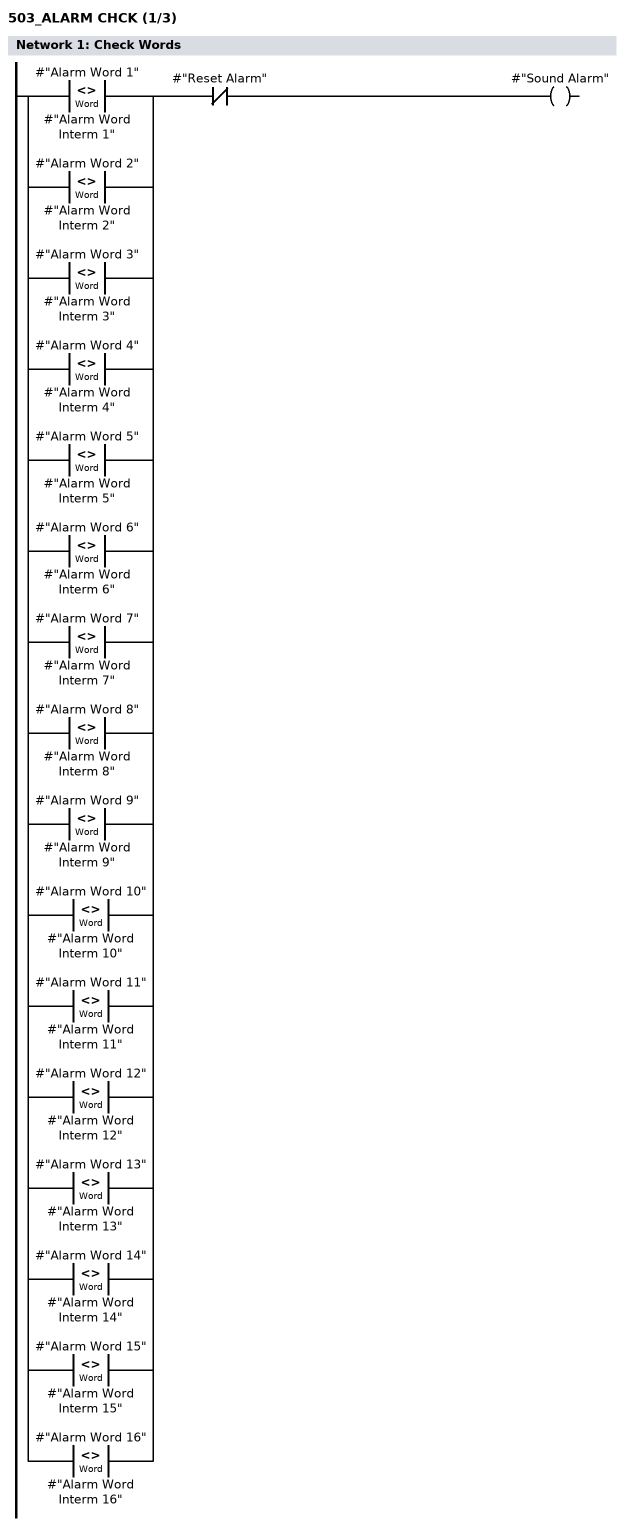
   RUNG wire#powerrail
      { S7_Templates := "SrcType := Word" } NE_Contact(in1 := #"Alarm Word 1", in2 := #"Alarm Word Interm 1")
      wire#w1
      I_Contact( #"Reset Alarm" )
      Coil( #"Sound Alarm" )
   END_RUNG
   RUNG wire#powerrail
      { S7_Templates := "SrcType := Word" } NE_Contact(in1 := #"Alarm Word 2", in2 := #"Alarm Word Interm 2")
   END_RUNG wire#w1
   RUNG wire#powerrail
      { S7_Templates := "SrcType := Word" } NE_Contact(in1 := #"Alarm Word 3", in2 := #"Alarm Word Interm 3")
   END_RUNG wire#w1
   RUNG wire#powerrail
      { S7_Templates := "SrcType := Word" } NE_Contact(in1 := #"Alarm Word 4", in2 := #"Alarm Word Interm 4")
   END_RUNG wire#w1
   RUNG wire#powerrail
      { S7_Templates := "SrcType := Word" } NE_Contact(in1 := #"Alarm Word 5", in2 := #"Alarm Word Interm 5")
   END_RUNG wire#w1
   RUNG wire#powerrail
      { S7_Templates := "SrcType := Word" } NE_Contact(in1 := #"Alarm Word 6", in2 := #"Alarm Word Interm 6")
   END_RUNG wire#w1
   RUNG wire#powerrail
      { S7_Templates := "SrcType := Word" } NE_Contact(in1 := #"Alarm Word 7", in2 := #"Alarm Word Interm 7")
   END_RUNG wire#w1
   RUNG wire#powerrail
      { S7_Templates := "SrcType := Word" } NE_Contact(in1 := #"Alarm Word 8", in2 := #"Alarm Word Interm 8")
   END_RUNG wire#w1
   RUNG wire#powerrail
      { S7_Templates := "SrcType := Word" } NE_Contact(in1 := #"Alarm Word 9", in2 := #"Alarm Word Interm 9")
   END_RUNG wire#w1
   RUNG wire#powerrail
      { S7_Templates := "SrcType := Word" } NE_Contact(in1 := #"Alarm Word 10", in2 := #"Alarm Word Interm 10")
   END_RUNG wire#w1
   RUNG wire#powerrail
      { S7_Templates := "SrcType := Word" } NE_Contact(in1 := #"Alarm Word 11", in2 := #"Alarm Word Interm 11")
   END_RUNG wire#w1
   RUNG wire#powerrail
      { S7_Templates := "SrcType := Word" } NE_Contact(in1 := #"Alarm Word 12", in2 := #"Alarm Word Interm 12")
   END_RUNG wire#w1
   RUNG wire#powerrail
      { S7_Templates := "SrcType := Word" } NE_Contact(in1 := #"Alarm Word 13", in2 := #"Alarm Word Interm 13")
   END_RUNG wire#w1
   RUNG wire#powerrail
      { S7_Templates := "SrcType := Word" } NE_Contact(in1 := #"Alarm Word 14", in2 := #"Alarm Word Interm 14")
   END_RUNG wire#w1
   RUNG wire#powerrail
      { S7_Templates := "SrcType := Word" } NE_Contact(in1 := #"Alarm Word 15", in2 := #"Alarm Word Interm 15")
   END_RUNG wire#w1
   RUNG wire#powerrail
      { S7_Templates := "SrcType := Word" } NE_Contact(in1 := #"Alarm Word 16", in2 := #"Alarm Word Interm 16")
   END_RUNG wire#w1
   // the same network as SCL:
   #"Sound Alarm" := ((#"Alarm Word 1" <> #"Alarm Word Interm 1") OR (#"Alarm Word 2" <> #"Alarm Word Interm 2") OR (#"Alarm Word 3" <> #"Alarm Word Interm 3") OR (#"Alarm Word 4" <> #"Alarm Word Interm 4") OR (#"Alarm Word 5" <> #"Alarm Word Interm 5") OR (#"Alarm Word 6" <> #"Alarm Word Interm 6") OR (#"Alarm Word 7" <> #"Alarm Word Interm 7") OR (#"Alarm Word 8" <> #"Alarm Word Interm 8") OR (#"Alarm Word 9" <> #"Alarm Word Interm 9") OR (#"Alarm Word 10" <> #"Alarm Word Interm 10") OR (#"Alarm Word 11" <> #"Alarm Word Interm 11") OR (#"Alarm Word 12" <> #"Alarm Word Interm 12") OR (#"Alarm Word 13" <> #"Alarm Word Interm 13") OR (#"Alarm Word 14" <> #"Alarm Word Interm 14") OR (#"Alarm Word 15" <> #"Alarm Word Interm 15") OR (#"Alarm Word 16" <> #"Alarm Word Interm 16")) AND NOT #"Reset Alarm";
END_REGION

REGION Network 2
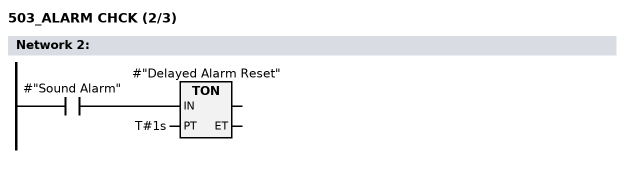
   #"Delayed Alarm Reset"(IN := #"Sound Alarm", PT := T#1s);   // TON
END_REGION

REGION Network 3: Move Words
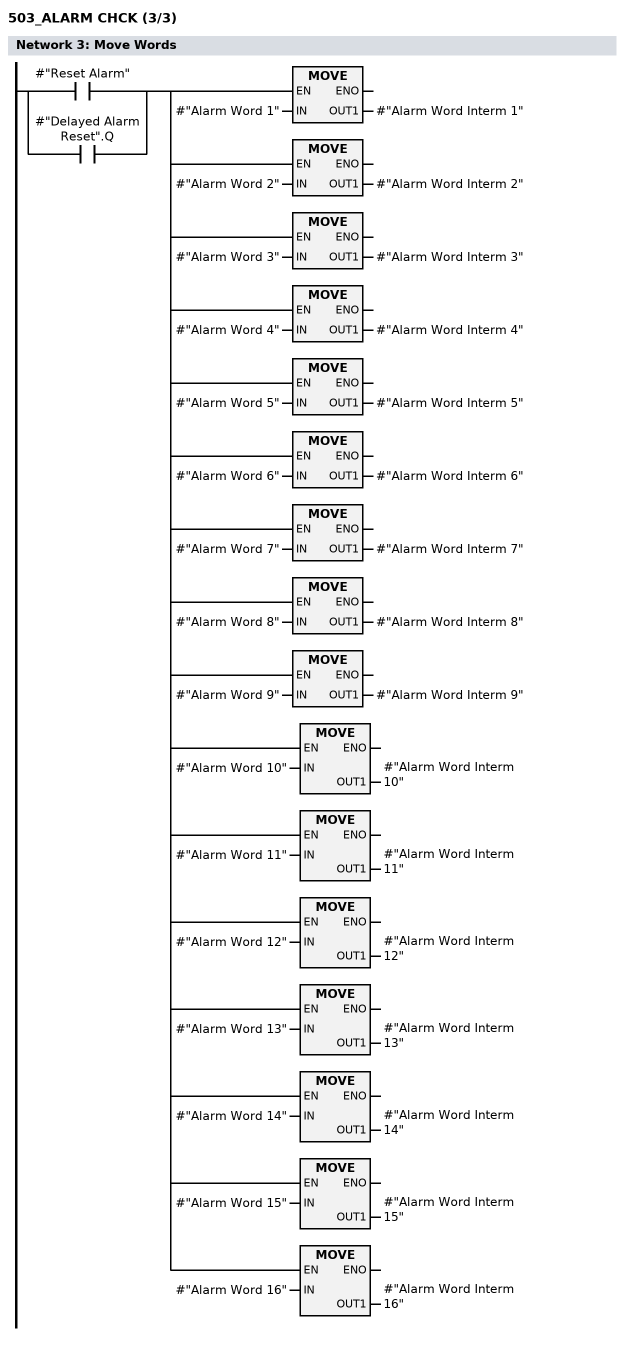
   RUNG wire#powerrail
      Contact( #"Reset Alarm" )
      wire#w1
      Move(in := #"Alarm Word 1", out1 => #"Alarm Word Interm 1")
   END_RUNG
   RUNG wire#powerrail
      Contact( #"Delayed Alarm Reset".Q )
   END_RUNG wire#w1
   RUNG wire#w1
      Move(in := #"Alarm Word 2", out1 => #"Alarm Word Interm 2")
   END_RUNG
   RUNG wire#w1
      Move(in := #"Alarm Word 3", out1 => #"Alarm Word Interm 3")
   END_RUNG
   RUNG wire#w1
      Move(in := #"Alarm Word 4", out1 => #"Alarm Word Interm 4")
   END_RUNG
   RUNG wire#w1
      Move(in := #"Alarm Word 5", out1 => #"Alarm Word Interm 5")
   END_RUNG
   RUNG wire#w1
      Move(in := #"Alarm Word 6", out1 => #"Alarm Word Interm 6")
   END_RUNG
   RUNG wire#w1
      Move(in := #"Alarm Word 7", out1 => #"Alarm Word Interm 7")
   END_RUNG
   RUNG wire#w1
      Move(in := #"Alarm Word 8", out1 => #"Alarm Word Interm 8")
   END_RUNG
   RUNG wire#w1
      Move(in := #"Alarm Word 9", out1 => #"Alarm Word Interm 9")
   END_RUNG
   RUNG wire#w1
      Move(in := #"Alarm Word 10", out1 => #"Alarm Word Interm 10")
   END_RUNG
   RUNG wire#w1
      Move(in := #"Alarm Word 11", out1 => #"Alarm Word Interm 11")
   END_RUNG
   RUNG wire#w1
      Move(in := #"Alarm Word 12", out1 => #"Alarm Word Interm 12")
   END_RUNG
   RUNG wire#w1
      Move(in := #"Alarm Word 13", out1 => #"Alarm Word Interm 13")
   END_RUNG
   RUNG wire#w1
      Move(in := #"Alarm Word 14", out1 => #"Alarm Word Interm 14")
   END_RUNG
   RUNG wire#w1
      Move(in := #"Alarm Word 15", out1 => #"Alarm Word Interm 15")
   END_RUNG
   RUNG wire#w1
      Move(in := #"Alarm Word 16", out1 => #"Alarm Word Interm 16")
   END_RUNG
   // the same network as SCL:
   IF #"Reset Alarm" OR #"Delayed Alarm Reset".Q THEN
       #"Alarm Word Interm 1" := #"Alarm Word 1";
       #"Alarm Word Interm 2" := #"Alarm Word 2";
       #"Alarm Word Interm 3" := #"Alarm Word 3";
       #"Alarm Word Interm 4" := #"Alarm Word 4";
       #"Alarm Word Interm 5" := #"Alarm Word 5";
       #"Alarm Word Interm 6" := #"Alarm Word 6";
       #"Alarm Word Interm 7" := #"Alarm Word 7";
       #"Alarm Word Interm 8" := #"Alarm Word 8";
       #"Alarm Word Interm 9" := #"Alarm Word 9";
       #"Alarm Word Interm 10" := #"Alarm Word 10";
       #"Alarm Word Interm 11" := #"Alarm Word 11";
       #"Alarm Word Interm 12" := #"Alarm Word 12";
       #"Alarm Word Interm 13" := #"Alarm Word 13";
       #"Alarm Word Interm 14" := #"Alarm Word 14";
       #"Alarm Word Interm 15" := #"Alarm Word 15";
       #"Alarm Word Interm 16" := #"Alarm Word 16";
   END_IF;
END_REGION
END_FUNCTION_BLOCK

FUNCTION_BLOCK "Choose"   // FB509, LAD
{ S7_Optimized_Access := 'TRUE' }
VERSION : 0.1
   VAR_INPUT
      Choose : Bool;
      "Option 1" : DInt;
      "Option 2" : DInt;
   END_VAR
   VAR_OUTPUT
      Output : DInt;
   END_VAR
   VAR
      True : Bool;
      False : Bool;
      "Option 1 M" : DInt;
      "Option 2 M" : DInt;
      "Choose Internal" : Bool;
      "Puls Aux" : Struct
         "Puls Aux 1" : Bool;
         "Puls Aux 2" : Bool;
         "Puls Aux 3" : Bool;
         "Puls Aux 4" : Bool;
         "Puls Aux 5" : Bool;
         "Puls Aux 6" : Bool;
      END_STRUCT;
      "TP P CHOOSE1" : TP_TIME;
      "TP N CHOOSE2" : TP_TIME;
      "TP N CHOOSE1" : TP_TIME;
      "TP P CHOOSE2" : TP_TIME;
      R_TRIG_Instance : R_TRIG;
      Puls : TP_TIME;
   END_VAR
   VAR_TEMP   // added for the SCL form of the ladder/FBD networks
      _w1 : Bool;
      _w2 : Bool;
      _w3 : Bool;
      _w4 : Bool;
   END_VAR
BEGIN

REGION Network 1: False/True
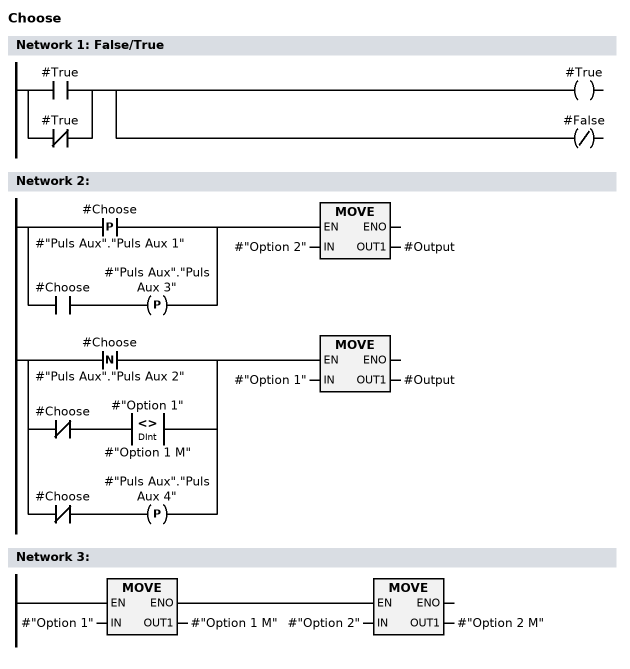
   RUNG wire#powerrail
      Contact( #True )
      wire#w1
      Coil( #True )
   END_RUNG
   RUNG wire#powerrail
      I_Contact( #True )
   END_RUNG wire#w1
   RUNG wire#w1
      I_Coil( #False )
   END_RUNG
   // the same network as SCL:
   #True := #True OR NOT #True;
   #False := NOT #True;
END_REGION

REGION Network 2
   RUNG wire#powerrail
      P_Contact(operand := #Choose, bit := #"Puls Aux"."Puls Aux 1")
      wire#w1
      Move(in := #"Option 2", out1 => #Output)
   END_RUNG
   RUNG wire#powerrail
      Contact( #Choose )
      P_Trig( #"Puls Aux"."Puls Aux 3" )
   END_RUNG wire#w1
   RUNG wire#powerrail
      N_Contact(operand := #Choose, bit := #"Puls Aux"."Puls Aux 2")
      wire#w2
      Move(in := #"Option 1", out1 => #Output)
   END_RUNG
   RUNG wire#powerrail
      I_Contact( #Choose )
      { S7_Templates := "SrcType := DInt" } NE_Contact(in1 := #"Option 1", in2 := #"Option 1 M")
   END_RUNG wire#w2
   RUNG wire#powerrail
      I_Contact( #Choose )
      P_Trig( #"Puls Aux"."Puls Aux 4" )
   END_RUNG wire#w2
   // the same network as SCL:
   #_w1 := #Choose AND NOT #"Puls Aux"."Puls Aux 1";   // rising edge of #Choose
   #"Puls Aux"."Puls Aux 1" := #Choose;
   #_w2 := #Choose AND NOT #"Puls Aux"."Puls Aux 3";   // rising edge
   #"Puls Aux"."Puls Aux 3" := #Choose;
   IF #_w1 OR #_w2 THEN #Output := #"Option 2"; END_IF;
   #_w3 := NOT #Choose AND #"Puls Aux"."Puls Aux 2";   // falling edge of #Choose
   #"Puls Aux"."Puls Aux 2" := #Choose;
   #_w4 := NOT #Choose AND NOT #"Puls Aux"."Puls Aux 4";   // rising edge
   #"Puls Aux"."Puls Aux 4" := NOT #Choose;
   IF #_w3 OR (NOT #Choose AND (#"Option 1" <> #"Option 1 M")) OR #_w4 THEN #Output := #"Option 1"; END_IF;
END_REGION

REGION Network 3
   RUNG wire#powerrail
      Move(in := #"Option 1", out1 => #"Option 1 M")
      Move(in := #"Option 2", out1 => #"Option 2 M")
   END_RUNG
   // the same network as SCL:
   #"Option 1 M" := #"Option 1";
   #"Option 2 M" := #"Option 2";
END_REGION
END_FUNCTION_BLOCK

FUNCTION_BLOCK "Flip Flop"   // FB510, LAD
{ S7_Optimized_Access := 'TRUE' }
VERSION : 0.1
   VAR_INPUT
      Input : Bool;
   END_VAR
   VAR_OUTPUT
      Output : Bool;
   END_VAR
   VAR
      SetOutputFlag : Bool;
   END_VAR
   VAR_TEMP   // added for the SCL form of the ladder/FBD networks
      _w1 : Bool;
      _w2 : Bool;
   END_VAR
BEGIN

REGION Network 2: Set Group SR
   // HMI Button to be set as SetTagWhileKeyPres
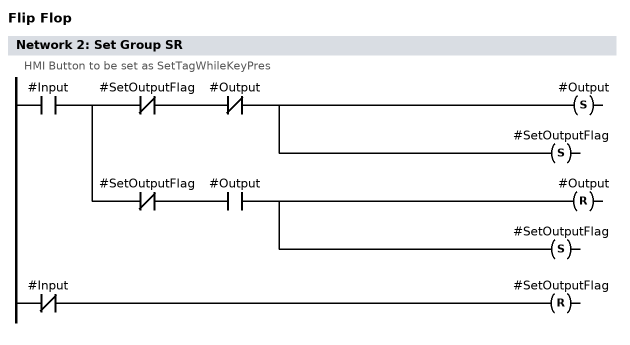
   RUNG wire#powerrail
      Contact( #Input )
      wire#w1
      I_Contact( #SetOutputFlag )
      I_Contact( #Output )
      wire#w2
      S_Coil( #Output )
   END_RUNG
   RUNG wire#w2
      S_Coil( #SetOutputFlag )
   END_RUNG
   RUNG wire#w1
      I_Contact( #SetOutputFlag )
      Contact( #Output )
      wire#w3
      R_Coil( #Output )
   END_RUNG
   RUNG wire#w3
      S_Coil( #SetOutputFlag )
   END_RUNG
   RUNG wire#powerrail
      I_Contact( #Input )
      R_Coil( #SetOutputFlag )
   END_RUNG
   // the same network as SCL:
   #_w1 := #Input AND NOT #SetOutputFlag AND NOT #Output;
   IF #_w1 THEN
       #Output := TRUE;
       #SetOutputFlag := TRUE;
   END_IF;
   #_w2 := #Input AND NOT #SetOutputFlag AND #Output;
   IF #_w2 THEN
       #Output := FALSE;
       #SetOutputFlag := TRUE;
   END_IF;
   IF NOT #Input THEN #SetOutputFlag := FALSE; END_IF;
END_REGION
END_FUNCTION_BLOCK

FUNCTION_BLOCK "Memory"   // FB511, LAD
{ S7_Optimized_Access := 'TRUE' }
VERSION : 0.1
   VAR_INPUT
      Enable : Bool;
      Negated : Bool := true;
      "Memorise/Remember" : Bool;
      Value : Int;
   END_VAR
   VAR_OUTPUT
      Remember : Int;
   END_VAR
   VAR RETAIN
      Memory : Int;
   END_VAR
   VAR
      PulsAuxP : Bool;
      PulsAuxN : Bool;
      SetOutputFlag : Bool;
      Output : Bool;
   END_VAR
   VAR_TEMP   // added for the SCL form of the ladder/FBD networks
      _w1 : Bool;
      _w2 : Bool;
      _w3 : Bool;
   END_VAR
BEGIN

REGION Network 1: Set Group SR
   // HMI Button to be set as SetTagWhileKeyPres
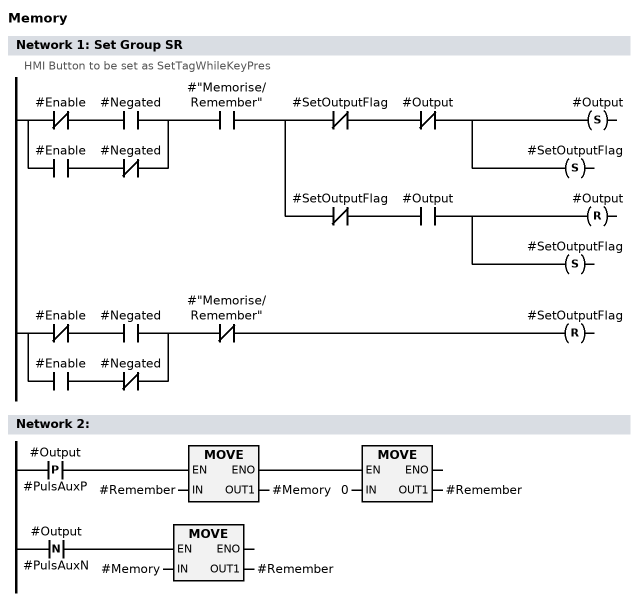
   RUNG wire#powerrail
      I_Contact( #Enable )
      Contact( #Negated )
      wire#w1
      Contact( #"Memorise/Remember" )
      wire#w2
      I_Contact( #SetOutputFlag )
      I_Contact( #Output )
      wire#w3
      S_Coil( #Output )
   END_RUNG
   RUNG wire#powerrail
      Contact( #Enable )
      I_Contact( #Negated )
   END_RUNG wire#w1
   RUNG wire#w3
      S_Coil( #SetOutputFlag )
   END_RUNG
   RUNG wire#w2
      I_Contact( #SetOutputFlag )
      Contact( #Output )
      wire#w4
      R_Coil( #Output )
   END_RUNG
   RUNG wire#w4
      S_Coil( #SetOutputFlag )
   END_RUNG
   RUNG wire#powerrail
      I_Contact( #Enable )
      Contact( #Negated )
      wire#w5
      I_Contact( #"Memorise/Remember" )
      R_Coil( #SetOutputFlag )
   END_RUNG
   RUNG wire#powerrail
      Contact( #Enable )
      I_Contact( #Negated )
   END_RUNG wire#w5
   // the same network as SCL:
   #_w1 := ((NOT #Enable AND #Negated) OR (#Enable AND NOT #Negated)) AND #"Memorise/Remember";
   #_w2 := #_w1 AND NOT #SetOutputFlag AND NOT #Output;
   IF #_w2 THEN
       #Output := TRUE;
       #SetOutputFlag := TRUE;
   END_IF;
   #_w3 := #_w1 AND NOT #SetOutputFlag AND #Output;
   IF #_w3 THEN
       #Output := FALSE;
       #SetOutputFlag := TRUE;
   END_IF;
   IF ((NOT #Enable AND #Negated) OR (#Enable AND NOT #Negated)) AND NOT #"Memorise/Remember" THEN
       #SetOutputFlag := FALSE;
   END_IF;
END_REGION

REGION Network 2
   RUNG wire#powerrail
      P_Contact(operand := #Output, bit := #PulsAuxP)
      Move(in := #Remember, out1 => #Memory)
      Move(in := 0, out1 => #Remember)
   END_RUNG
   RUNG wire#powerrail
      N_Contact(operand := #Output, bit := #PulsAuxN)
      Move(in := #Memory, out1 => #Remember)
   END_RUNG
   // the same network as SCL:
   #_w1 := #Output AND NOT #PulsAuxP;   // rising edge of #Output
   #PulsAuxP := #Output;
   IF #_w1 THEN
       #Memory := #Remember;
       #Remember := 0;
   END_IF;
   #_w2 := NOT #Output AND #PulsAuxN;   // falling edge of #Output
   #PulsAuxN := #Output;
   IF #_w2 THEN #Remember := #Memory; END_IF;
END_REGION
END_FUNCTION_BLOCK

FUNCTION_BLOCK "Sequence Times"   // FB512, LAD
{ S7_Optimized_Access := 'TRUE' }
VERSION : 0.1
   VAR_INPUT
      "Start Jurney" : Bool;
      "Start De-Ox" : Bool;
      "Start Dwell" : Bool;
      "Start Re-Ox" : Bool;
      "Start Post-Dwell" : Bool;
      "Jurney Time" : Real := 30.0;   // Days
      "Pre-Dwell Time" : Real := 1.0;   // Hours
      "De-Ox Time" : Real := 12.0;   // Hours
      "De-Ox SP Time" : Real := 1.0;   // Hours
      "De-Ox O2 Confirm" : Real := 1.0;   // Minutes
      "Dwell Time" : Real := 60.0;   // Hours
      "Re-Ox Time" : Real := 6.0;   // Hours
      "Post-Dwell Time" : Real := 12.0;   // Hours
      "Offset Treatment Time" : Real := 0.0;   // Hours
      "Offset Treatment Time Extend" : Real := 13.0;
      "Offset De-Ox Time Extend" : Real;
      "Offset Re-Ox Time Extend" : Real;
      "Time to IGG Start Warning" : DInt;   // Hours
      Continue : Bool;
      Boost : Bool;
   END_VAR
   VAR_OUTPUT
      "Times Valid" : Bool;
      "Warn to IGG Start" : Bool;
      "Warn to GCU Start" : Bool;   // Warning to start GCU at Re-Ox
      "Pre-Dwell Done" : Bool;
      "De-Ox Done" : Bool;
      "Dwell Done" : Bool;
      "Re-Ox Done" : Bool;
      "Post-Dwell Done" : Bool;
      "Pre-Dwell Time Corected" : Real;
      "Voiage Time Invalid" : Bool;
   END_VAR
   VAR
      "Extra Time" : Real;
      "Jurney Aux" : Time;
      "Pre-Dwell Aux" : Real;
      "Pre-Dwell Aux Memory" : Real;
   END_VAR
   VAR RETAIN
      "Pre-Dwell Memory h" : Real;
   END_VAR
   VAR
      "De-Ox Aux" : Real;
      "De-Ox Aux Memory" : Real;
   END_VAR
   VAR RETAIN
      "De-Ox Memory h" : Real;
   END_VAR
   VAR
      "Dwell Aux" : Real;
      "Dwell Aux Memory" : Real;
   END_VAR
   VAR RETAIN
      "Dwell Memory h" : Real;
   END_VAR
   VAR
      "Re-Ox Aux" : Real;
      "Re-Ox Aux Memory" : Real;
   END_VAR
   VAR RETAIN
      "Re-Ox Memory h" : Real;
   END_VAR
   VAR
      "Post-Dwell Aux" : Real;
      "Post-Dwell Aux Memory" : Real;
   END_VAR
   VAR RETAIN
      "Post-Dwell Memory h" : Real;
   END_VAR
   VAR
      True : Bool;
      False : Bool;
      "Pulse Continue" : Bool;
      IEC_Timer_0_Instance : TON_TIME;
      "Jurney Time FB" : "Days Timer";
      "Pre-Dwell Timer" : "Hours Timer";
      "Dwell Timer" : "Hours Timer";
      "Post-Dwell Timer" : "Hours Timer";
      "Puls Timer" : TON_TIME;
      "Puls TP" : TP_TIME;
      "Treatment Timer" : "Hours Timer";
      "De-Ox Timer" : "Hours Timer";
      "Re-Ox Timer" : "Hours Timer";
      "Jurney Timer" : "Hours Timer";
      "Offset Timer" : "Hours Timer";
      "Flip Flop_Pre-Dwell" : "Flip Flop";
      "Choose_Instance_Pre-Dwell" : "Choose Real";
      "Choose_Instance_De-Ox" : "Choose Real";
      Choose_Instance_Dwell : "Choose Real";
      "Choose_Instance_Re-Ox" : "Choose Real";
      "Choose_Instance_Post-Dwell" : "Choose Real";
   END_VAR
   VAR_TEMP   // added for the SCL form of the ladder/FBD networks
      _w1 : Bool;
   END_VAR
BEGIN

REGION Network 1
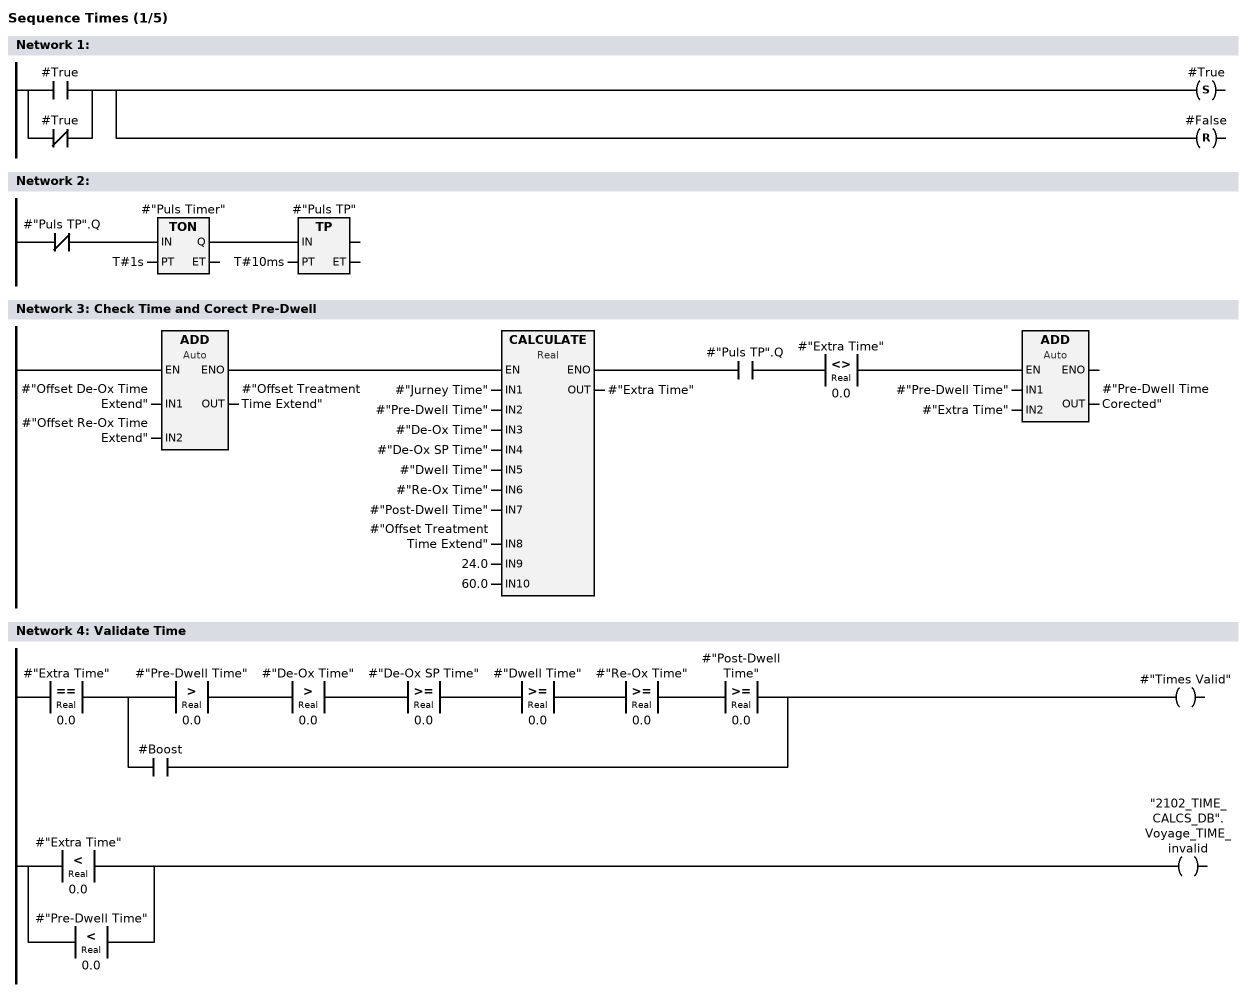
   RUNG wire#powerrail
      Contact( #True )
      wire#w1
      S_Coil( #True )
   END_RUNG
   RUNG wire#powerrail
      I_Contact( #True )
   END_RUNG wire#w1
   RUNG wire#w1
      R_Coil( #False )
   END_RUNG
   // the same network as SCL:
   #_w1 := #True OR NOT #True;
   IF #_w1 THEN
       #True := TRUE;
       #False := FALSE;
   END_IF;
END_REGION

REGION Network 2
   #"Puls Timer"(IN := NOT #"Puls TP".Q, PT := T#1s);   // TON
   #"Puls TP"(IN := #"Puls Timer".Q, PT := T#10ms);   // TP
END_REGION

REGION Network 3: Check Time and Corect Pre-Dwell
   RUNG wire#powerrail
      Add(in1 := #"Offset De-Ox Time Extend", in2 := #"Offset Re-Ox Time Extend", out => #"Offset Treatment Time Extend")
      { S7_Templates := "SrcType := Real"; S7_Expression := "IN1*IN9-(IN2+IN3+IN4+IN5+IN6+IN7+IN8)" } Calculate(in1 := #"Jurney Time", in2 := #"Pre-Dwell Time", in3 := #"De-Ox Time", in4 := #"De-Ox SP Time", in5 := #"Dwell Time", in6 := #"Re-Ox Time", in7 := #"Post-Dwell Time", in8 := #"Offset Treatment Time Extend", in9 := 24.0, in10 := 60.0, out => #"Extra Time")
      Contact( #"Puls TP".Q )
      { S7_Templates := "SrcType := Real" } NE_Contact(in1 := #"Extra Time", in2 := 0.0)
      Add(in1 := #"Pre-Dwell Time", in2 := #"Extra Time", out => #"Pre-Dwell Time Corected")
   END_RUNG
   // the same network as SCL:
   #"Offset Treatment Time Extend" := #"Offset De-Ox Time Extend" + #"Offset Re-Ox Time Extend";
   #"Extra Time" := #"Jurney Time"*24.0-(#"Pre-Dwell Time"+#"De-Ox Time"+#"De-Ox SP Time"+#"Dwell Time"+#"Re-Ox Time"+#"Post-Dwell Time"+#"Offset Treatment Time Extend");
   IF #"Puls TP".Q AND (#"Extra Time" <> 0.0) THEN
       #"Pre-Dwell Time Corected" := #"Pre-Dwell Time" + #"Extra Time";
   END_IF;
END_REGION

REGION Network 4: Validate Time
   RUNG wire#powerrail
      { S7_Templates := "SrcType := Real" } EQ_Contact(in1 := #"Extra Time", in2 := 0.0)
      wire#w1
      { S7_Templates := "SrcType := Real" } GT_Contact(in1 := #"Pre-Dwell Time", in2 := 0.0)
      { S7_Templates := "SrcType := Real" } GT_Contact(in1 := #"De-Ox Time", in2 := 0.0)
      { S7_Templates := "SrcType := Real" } GE_Contact(in1 := #"De-Ox SP Time", in2 := 0.0)
      { S7_Templates := "SrcType := Real" } GE_Contact(in1 := #"Dwell Time", in2 := 0.0)
      { S7_Templates := "SrcType := Real" } GE_Contact(in1 := #"Re-Ox Time", in2 := 0.0)
      { S7_Templates := "SrcType := Real" } GE_Contact(in1 := #"Post-Dwell Time", in2 := 0.0)
      wire#w2
      Coil( #"Times Valid" )
   END_RUNG
   RUNG wire#w1
      Contact( #Boost )
   END_RUNG wire#w2
   RUNG wire#powerrail
      { S7_Templates := "SrcType := Real" } LT_Contact(in1 := #"Extra Time", in2 := 0.0)
      wire#w3
      Coil( "2102_TIME_CALCS_DB".Voyage_TIME_invalid )
   END_RUNG
   RUNG wire#powerrail
      { S7_Templates := "SrcType := Real" } LT_Contact(in1 := #"Pre-Dwell Time", in2 := 0.0)
   END_RUNG wire#w3
   // the same network as SCL:
   #"Times Valid" := (#"Extra Time" = 0.0) AND (((#"Pre-Dwell Time" > 0.0) AND (#"De-Ox Time" > 0.0) AND (#"De-Ox SP Time" >= 0.0) AND (#"Dwell Time" >= 0.0) AND (#"Re-Ox Time" >= 0.0) AND (#"Post-Dwell Time" >= 0.0)) OR #Boost);
   "2102_TIME_CALCS_DB".Voyage_TIME_invalid := (#"Extra Time" < 0.0) OR (#"Pre-Dwell Time" < 0.0);
END_REGION

REGION Network 5: Total Sequence Time
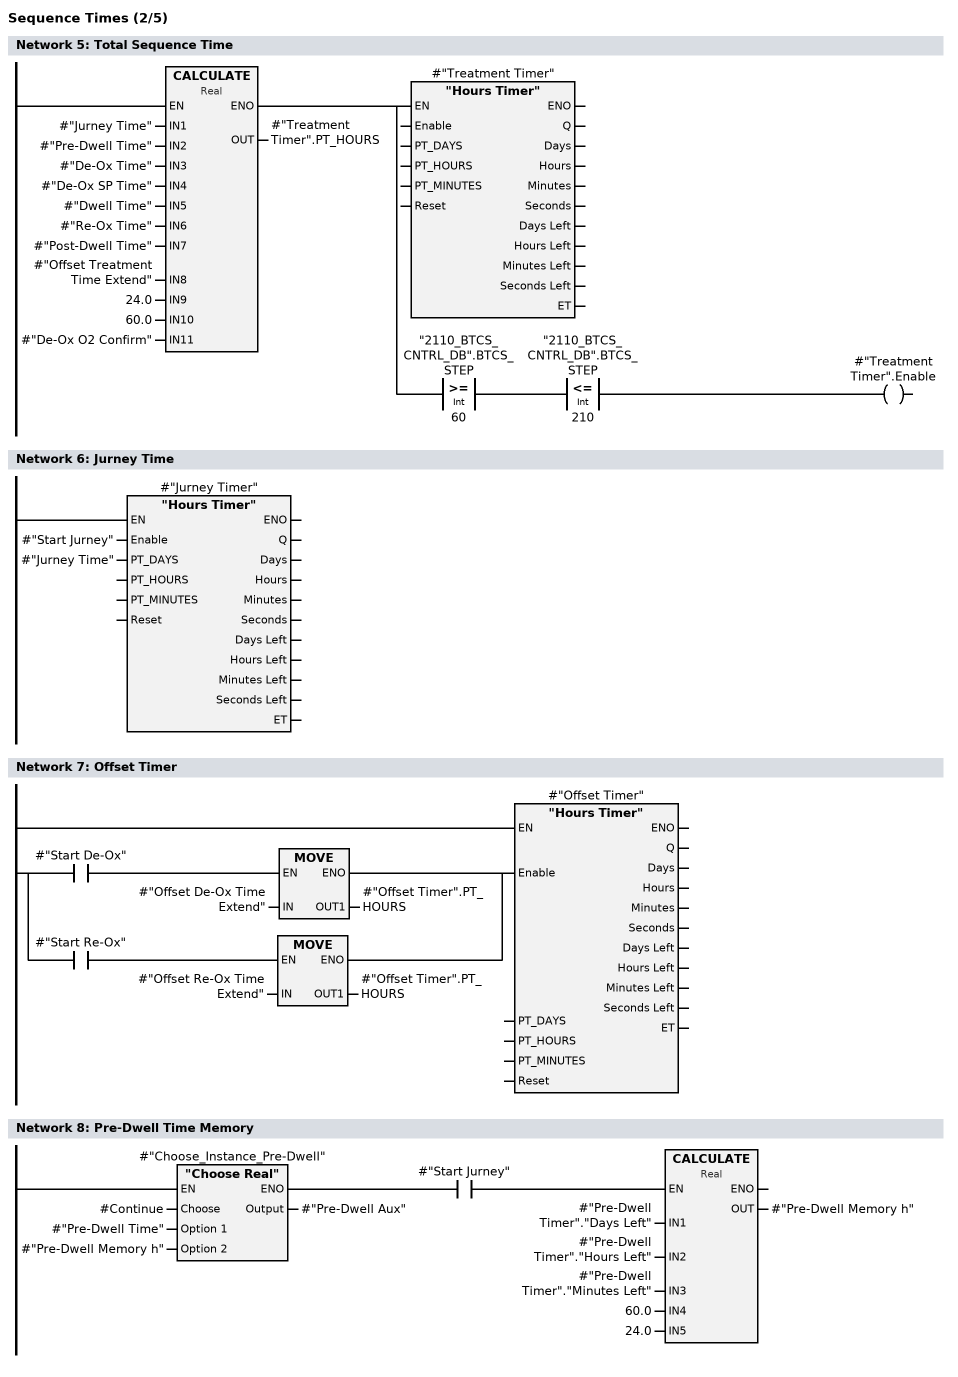
   RUNG wire#powerrail
      { S7_Templates := "SrcType := Real"; S7_Expression := "IN3+IN4+IN5+IN6+IN7+IN8+(IN11/IN10)" } Calculate(in1 := #"Jurney Time", in2 := #"Pre-Dwell Time", in3 := #"De-Ox Time", in4 := #"De-Ox SP Time", in5 := #"Dwell Time", in6 := #"Re-Ox Time", in7 := #"Post-Dwell Time", in8 := #"Offset Treatment Time Extend", in9 := 24.0, in10 := 60.0, in11 := #"De-Ox O2 Confirm", out => #"Treatment Timer".PT_HOURS)
      wire#w1
      #"Treatment Timer"(Enable :=, PT_DAYS :=, PT_HOURS :=, PT_MINUTES :=, Reset :=, Q =>, Days =>, Hours =>, Minutes =>, Seconds =>, "Days Left" =>, "Hours Left" =>, "Minutes Left" =>, "Seconds Left" =>, ET =>)
   END_RUNG
   RUNG wire#w1
      { S7_Templates := "SrcType := Int" } GE_Contact(in1 := "2110_BTCS_CNTRL_DB".BTCS_STEP, in2 := 60)
      { S7_Templates := "SrcType := Int" } LE_Contact(in1 := "2110_BTCS_CNTRL_DB".BTCS_STEP, in2 := 210)
      Coil( #"Treatment Timer".Enable )
   END_RUNG
   // the same network as SCL:
   #"Treatment Timer".PT_HOURS := #"De-Ox Time"+#"De-Ox SP Time"+#"Dwell Time"+#"Re-Ox Time"+#"Post-Dwell Time"+#"Offset Treatment Time Extend"+(#"De-Ox O2 Confirm"/60.0);
   #"Treatment Timer"();   // "Hours Timer"
   #"Treatment Timer".Enable := ("2110_BTCS_CNTRL_DB".BTCS_STEP >= 60) AND ("2110_BTCS_CNTRL_DB".BTCS_STEP <= 210);
END_REGION

REGION Network 6: Jurney Time
   RUNG wire#powerrail
      #"Jurney Timer"(Enable := #"Start Jurney", PT_DAYS := #"Jurney Time", PT_HOURS :=, PT_MINUTES :=, Reset :=, Q =>, Days =>, Hours =>, Minutes =>, Seconds =>, "Days Left" =>, "Hours Left" =>, "Minutes Left" =>, "Seconds Left" =>, ET =>)
   END_RUNG
   // the same network as SCL:
   #"Jurney Timer"(Enable := #"Start Jurney", PT_DAYS := #"Jurney Time");   // "Hours Timer"
END_REGION

REGION Network 7: Offset Timer
   RUNG wire#powerrail
      #"Offset Timer"(Enable := wire#w1, PT_DAYS :=, PT_HOURS :=, PT_MINUTES :=, Reset :=, Q =>, Days =>, Hours =>, Minutes =>, Seconds =>, "Days Left" =>, "Hours Left" =>, "Minutes Left" =>, "Seconds Left" =>, ET =>)
   END_RUNG
   RUNG wire#powerrail
      Contact( #"Start De-Ox" )
      Move(in := #"Offset De-Ox Time Extend", out1 => #"Offset Timer".PT_HOURS)
   END_RUNG wire#w1
   RUNG wire#powerrail
      Contact( #"Start Re-Ox" )
      Move(in := #"Offset Re-Ox Time Extend", out1 => #"Offset Timer".PT_HOURS)
   END_RUNG wire#w1
   // the same network as SCL:
   IF #"Start De-Ox" THEN #"Offset Timer".PT_HOURS := #"Offset De-Ox Time Extend"; END_IF;
   IF #"Start Re-Ox" THEN #"Offset Timer".PT_HOURS := #"Offset Re-Ox Time Extend"; END_IF;
   #"Offset Timer"(Enable := #"Start De-Ox" OR #"Start Re-Ox");   // "Hours Timer"
END_REGION

REGION Network 8: Pre-Dwell Time Memory
   RUNG wire#powerrail
      #"Choose_Instance_Pre-Dwell"(Choose := #Continue, "Option 1" := #"Pre-Dwell Time", "Option 2" := #"Pre-Dwell Memory h", Output => #"Pre-Dwell Aux")
      Contact( #"Start Jurney" )
      { S7_Templates := "SrcType := Real"; S7_Expression := "(IN1*IN5)+IN2+(IN3/IN4)" } Calculate(in1 := #"Pre-Dwell Timer"."Days Left", in2 := #"Pre-Dwell Timer"."Hours Left", in3 := #"Pre-Dwell Timer"."Minutes Left", in4 := 60.0, in5 := 24.0, out => #"Pre-Dwell Memory h")
   END_RUNG
   // the same network as SCL:
   #"Choose_Instance_Pre-Dwell"(Choose := #Continue,   // "Choose Real"
                           "Option 1" := #"Pre-Dwell Time",
                           "Option 2" := #"Pre-Dwell Memory h",
                           Output => #"Pre-Dwell Aux",
                           ENO => #_w1);
   IF #_w1 AND #"Start Jurney" THEN
       #"Pre-Dwell Memory h" := (#"Pre-Dwell Timer"."Days Left"*24.0)+#"Pre-Dwell Timer"."Hours Left"+(#"Pre-Dwell Timer"."Minutes Left"/60.0);
   END_IF;
END_REGION

REGION Network 9: Pre-Dwell remaining
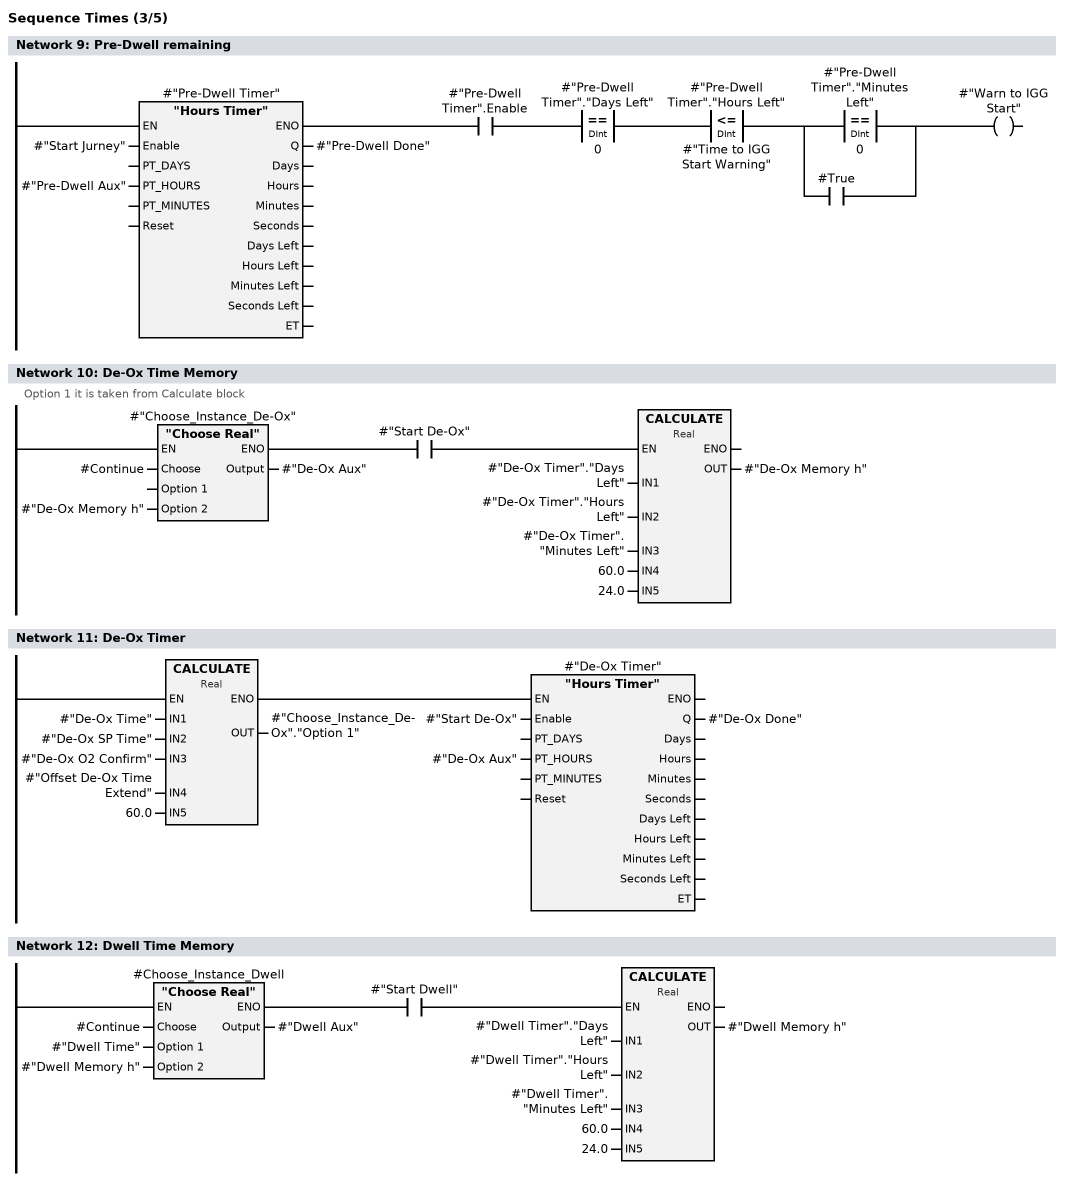
   RUNG wire#powerrail
      #"Pre-Dwell Timer"(Enable := #"Start Jurney", PT_DAYS :=, PT_HOURS := #"Pre-Dwell Aux", PT_MINUTES :=, Reset :=, Q => #"Pre-Dwell Done", Days =>, Hours =>, Minutes =>, Seconds =>, "Days Left" =>, "Hours Left" =>, "Minutes Left" =>, "Seconds Left" =>, ET =>)
      Contact( #"Pre-Dwell Timer".Enable )
      { S7_Templates := "SrcType := DInt" } EQ_Contact(in1 := #"Pre-Dwell Timer"."Days Left", in2 := 0)
      { S7_Templates := "SrcType := DInt" } LE_Contact(in1 := #"Pre-Dwell Timer"."Hours Left", in2 := #"Time to IGG Start Warning")
      wire#w1
      { S7_Templates := "SrcType := DInt" } EQ_Contact(in1 := #"Pre-Dwell Timer"."Minutes Left", in2 := 0)
      wire#w2
      Coil( #"Warn to IGG Start" )
   END_RUNG
   RUNG wire#w1
      Contact( #True )
   END_RUNG wire#w2
   // the same network as SCL:
   #"Pre-Dwell Timer"(Enable := #"Start Jurney",   // "Hours Timer"
                      PT_HOURS := #"Pre-Dwell Aux",
                      Q => #"Pre-Dwell Done",
                      ENO => #_w1);
   #"Warn to IGG Start" := #_w1 AND #"Pre-Dwell Timer".Enable AND (#"Pre-Dwell Timer"."Days Left" = 0) AND (#"Pre-Dwell Timer"."Hours Left" <= #"Time to IGG Start Warning") AND ((#"Pre-Dwell Timer"."Minutes Left" = 0) OR #True);
END_REGION

REGION Network 10: De-Ox Time Memory
   // Option 1 it is taken from Calculate block
   RUNG wire#powerrail
      #"Choose_Instance_De-Ox"(Choose := #Continue, "Option 1" :=, "Option 2" := #"De-Ox Memory h", Output => #"De-Ox Aux")
      Contact( #"Start De-Ox" )
      { S7_Templates := "SrcType := Real"; S7_Expression := "(IN1*IN5)+IN2+(IN3/IN4)" } Calculate(in1 := #"De-Ox Timer"."Days Left", in2 := #"De-Ox Timer"."Hours Left", in3 := #"De-Ox Timer"."Minutes Left", in4 := 60.0, in5 := 24.0, out => #"De-Ox Memory h")
   END_RUNG
   // the same network as SCL:
   #"Choose_Instance_De-Ox"(Choose := #Continue,   // "Choose Real"
                           "Option 2" := #"De-Ox Memory h",
                           Output => #"De-Ox Aux",
                           ENO => #_w1);
   IF #_w1 AND #"Start De-Ox" THEN
       #"De-Ox Memory h" := (#"De-Ox Timer"."Days Left"*24.0)+#"De-Ox Timer"."Hours Left"+(#"De-Ox Timer"."Minutes Left"/60.0);
   END_IF;
END_REGION

REGION Network 11: De-Ox Timer
   RUNG wire#powerrail
      { S7_Templates := "SrcType := Real"; S7_Expression := "IN1+IN2+(IN3/IN5)+IN4" } Calculate(in1 := #"De-Ox Time", in2 := #"De-Ox SP Time", in3 := #"De-Ox O2 Confirm", in4 := #"Offset De-Ox Time Extend", in5 := 60.0, out => #"Choose_Instance_De-Ox"."Option 1")
      #"De-Ox Timer"(Enable := #"Start De-Ox", PT_DAYS :=, PT_HOURS := #"De-Ox Aux", PT_MINUTES :=, Reset :=, Q => #"De-Ox Done", Days =>, Hours =>, Minutes =>, Seconds =>, "Days Left" =>, "Hours Left" =>, "Minutes Left" =>, "Seconds Left" =>, ET =>)
   END_RUNG
   // the same network as SCL:
   #"Choose_Instance_De-Ox"."Option 1" := #"De-Ox Time"+#"De-Ox SP Time"+(#"De-Ox O2 Confirm"/60.0)+#"Offset De-Ox Time Extend";
   #"De-Ox Timer"(Enable := #"Start De-Ox", PT_HOURS := #"De-Ox Aux", Q => #"De-Ox Done");   // "Hours Timer"
END_REGION

REGION Network 12: Dwell Time Memory
   RUNG wire#powerrail
      #Choose_Instance_Dwell(Choose := #Continue, "Option 1" := #"Dwell Time", "Option 2" := #"Dwell Memory h", Output => #"Dwell Aux")
      Contact( #"Start Dwell" )
      { S7_Templates := "SrcType := Real"; S7_Expression := "(IN1*IN5)+IN2+(IN3/IN4)" } Calculate(in1 := #"Dwell Timer"."Days Left", in2 := #"Dwell Timer"."Hours Left", in3 := #"Dwell Timer"."Minutes Left", in4 := 60.0, in5 := 24.0, out => #"Dwell Memory h")
   END_RUNG
   // the same network as SCL:
   #Choose_Instance_Dwell(Choose := #Continue,   // "Choose Real"
                          "Option 1" := #"Dwell Time",
                          "Option 2" := #"Dwell Memory h",
                          Output => #"Dwell Aux",
                          ENO => #_w1);
   IF #_w1 AND #"Start Dwell" THEN
       #"Dwell Memory h" := (#"Dwell Timer"."Days Left"*24.0)+#"Dwell Timer"."Hours Left"+(#"Dwell Timer"."Minutes Left"/60.0);
   END_IF;
END_REGION

REGION Network 13: Dwell Remaining
